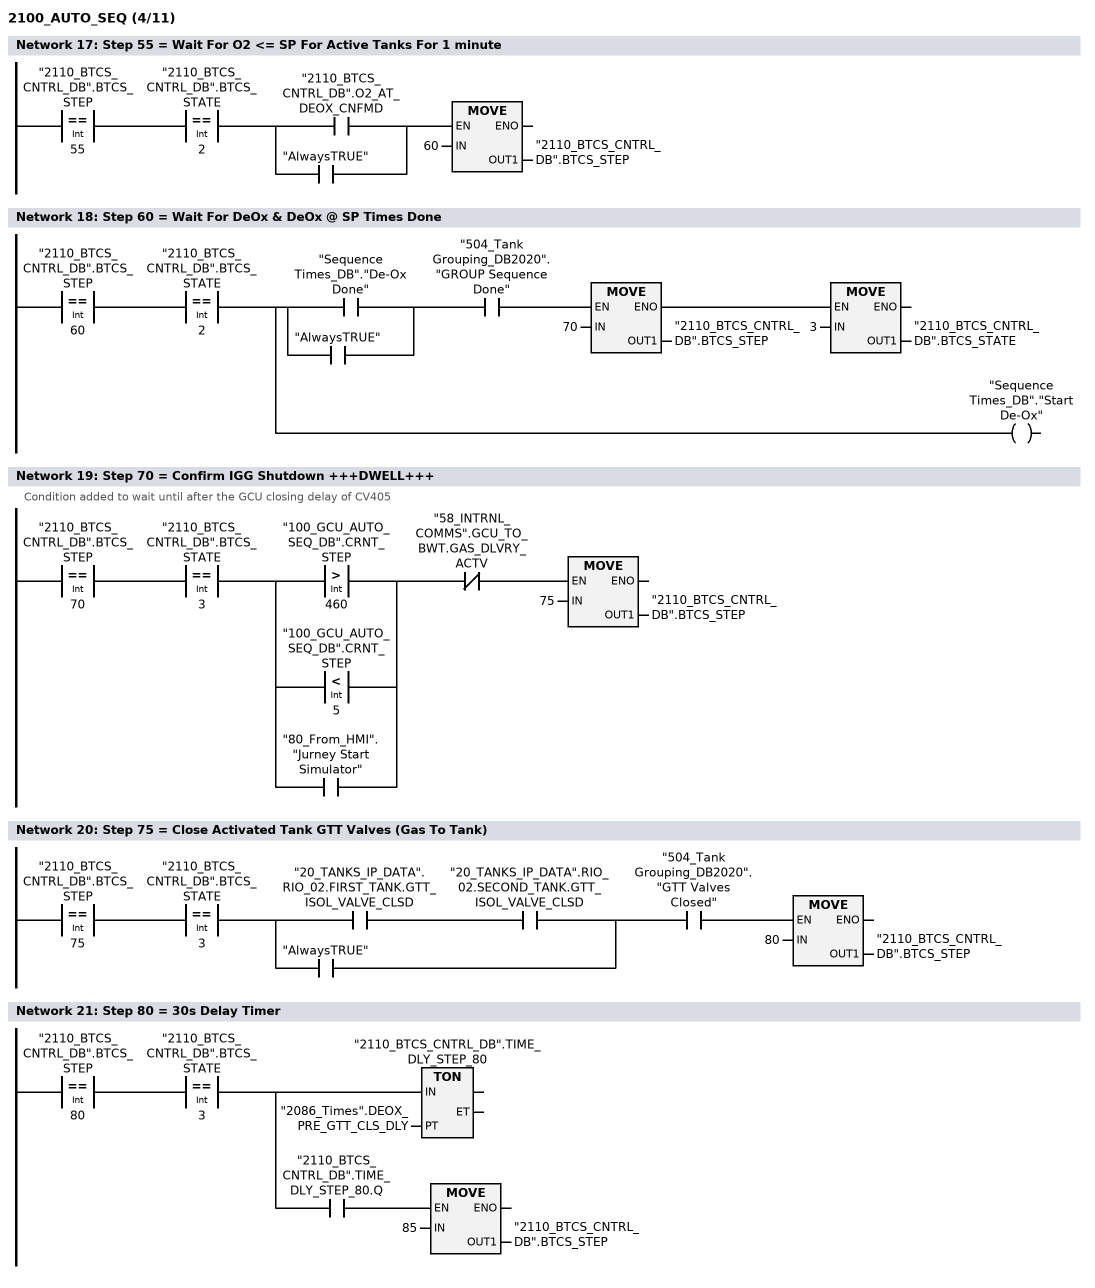
   RUNG wire#powerrail
      { S7_Templates := "SrcType := Int" } EQ_Contact(in1 := "2110_BTCS_CNTRL_DB".BTCS_STEP, in2 := 55)
      { S7_Templates := "SrcType := Int" } EQ_Contact(in1 := "2110_BTCS_CNTRL_DB".BTCS_STATE, in2 := 2)
      wire#w1
      Contact( "2110_BTCS_CNTRL_DB".O2_AT_DEOX_CNFMD )
      wire#w2
      Move(in := 60, out1 => "2110_BTCS_CNTRL_DB".BTCS_STEP)
   END_RUNG
   RUNG wire#w1
      Contact( "AlwaysTRUE" )
   END_RUNG wire#w2
   // the same network as SCL:
   IF ("2110_BTCS_CNTRL_DB".BTCS_STEP = 55) AND ("2110_BTCS_CNTRL_DB".BTCS_STATE = 2) AND ("2110_BTCS_CNTRL_DB".O2_AT_DEOX_CNFMD OR "AlwaysTRUE") THEN
       "2110_BTCS_CNTRL_DB".BTCS_STEP := 60;
   END_IF;
END_REGION

REGION Network 18: Step 60 = Wait For DeOx & DeOx @ SP Times Done
   RUNG wire#powerrail
      { S7_Templates := "SrcType := Int" } EQ_Contact(in1 := "2110_BTCS_CNTRL_DB".BTCS_STEP, in2 := 60)
      { S7_Templates := "SrcType := Int" } EQ_Contact(in1 := "2110_BTCS_CNTRL_DB".BTCS_STATE, in2 := 2)
      wire#w1
      Contact( "Sequence Times_DB"."De-Ox Done" )
      wire#w2
      Contact( "504_Tank Grouping_DB2020"."GROUP Sequence Done" )
      Move(in := 70, out1 => "2110_BTCS_CNTRL_DB".BTCS_STEP)
      Move(in := 3, out1 => "2110_BTCS_CNTRL_DB".BTCS_STATE)
   END_RUNG
   RUNG wire#w1
      Contact( "AlwaysTRUE" )
   END_RUNG wire#w2
   RUNG wire#w1
      Coil( "Sequence Times_DB"."Start De-Ox" )
   END_RUNG
   // the same network as SCL:
   #_w1 := ("2110_BTCS_CNTRL_DB".BTCS_STEP = 60) AND ("2110_BTCS_CNTRL_DB".BTCS_STATE = 2);
   IF #_w1 AND ("Sequence Times_DB"."De-Ox Done" OR "AlwaysTRUE") AND "504_Tank Grouping_DB2020"."GROUP Sequence Done" THEN
       "2110_BTCS_CNTRL_DB".BTCS_STEP := 70;
       "2110_BTCS_CNTRL_DB".BTCS_STATE := 3;
   END_IF;
   "Sequence Times_DB"."Start De-Ox" := #_w1;
END_REGION

REGION Network 19: Step 70 = Confirm IGG Shutdown +++DWELL+++
   // Condition added to wait until after the GCU closing delay of CV405
   RUNG wire#powerrail
      { S7_Templates := "SrcType := Int" } EQ_Contact(in1 := "2110_BTCS_CNTRL_DB".BTCS_STEP, in2 := 70)
      { S7_Templates := "SrcType := Int" } EQ_Contact(in1 := "2110_BTCS_CNTRL_DB".BTCS_STATE, in2 := 3)
      wire#w1
      { S7_Templates := "SrcType := Int" } GT_Contact(in1 := "100_GCU_AUTO_SEQ_DB".CRNT_STEP, in2 := 460)
      wire#w2
      I_Contact( "58_INTRNL_COMMS".GCU_TO_BWT.GAS_DLVRY_ACTV )
      Move(in := 75, out1 => "2110_BTCS_CNTRL_DB".BTCS_STEP)
   END_RUNG
   RUNG wire#w1
      { S7_Templates := "SrcType := Int" } LT_Contact(in1 := "100_GCU_AUTO_SEQ_DB".CRNT_STEP, in2 := 5)
   END_RUNG wire#w2
   RUNG wire#w1
      Contact( "80_From_HMI"."Jurney Start Simulator" )
   END_RUNG wire#w2
   // the same network as SCL:
   IF ("2110_BTCS_CNTRL_DB".BTCS_STEP = 70) AND ("2110_BTCS_CNTRL_DB".BTCS_STATE = 3) AND (("100_GCU_AUTO_SEQ_DB".CRNT_STEP > 460) OR ("100_GCU_AUTO_SEQ_DB".CRNT_STEP < 5) OR "80_From_HMI"."Jurney Start Simulator") AND NOT "58_INTRNL_COMMS".GCU_TO_BWT.GAS_DLVRY_ACTV THEN
       "2110_BTCS_CNTRL_DB".BTCS_STEP := 75;
   END_IF;
END_REGION

REGION Network 20: Step 75 = Close Activated Tank GTT Valves (Gas To Tank)
   RUNG wire#powerrail
      { S7_Templates := "SrcType := Int" } EQ_Contact(in1 := "2110_BTCS_CNTRL_DB".BTCS_STEP, in2 := 75)
      { S7_Templates := "SrcType := Int" } EQ_Contact(in1 := "2110_BTCS_CNTRL_DB".BTCS_STATE, in2 := 3)
      wire#w1
      Contact( "20_TANKS_IP_DATA".RIO_02.FIRST_TANK.GTT_ISOL_VALVE_CLSD )
      Contact( "20_TANKS_IP_DATA".RIO_02.SECOND_TANK.GTT_ISOL_VALVE_CLSD )
      wire#w2
      Contact( "504_Tank Grouping_DB2020"."GTT Valves Closed" )
      Move(in := 80, out1 => "2110_BTCS_CNTRL_DB".BTCS_STEP)
   END_RUNG
   RUNG wire#w1
      Contact( "AlwaysTRUE" )
   END_RUNG wire#w2
   // the same network as SCL:
   IF ("2110_BTCS_CNTRL_DB".BTCS_STEP = 75) AND ("2110_BTCS_CNTRL_DB".BTCS_STATE = 3) AND (("20_TANKS_IP_DATA".RIO_02.FIRST_TANK.GTT_ISOL_VALVE_CLSD AND "20_TANKS_IP_DATA".RIO_02.SECOND_TANK.GTT_ISOL_VALVE_CLSD) OR "AlwaysTRUE") AND "504_Tank Grouping_DB2020"."GTT Valves Closed" THEN
       "2110_BTCS_CNTRL_DB".BTCS_STEP := 80;
   END_IF;
END_REGION

REGION Network 21: Step 80 = 30s Delay Timer
   #_w1 := ("2110_BTCS_CNTRL_DB".BTCS_STEP = 80) AND ("2110_BTCS_CNTRL_DB".BTCS_STATE = 3);
   "2110_BTCS_CNTRL_DB".TIME_DLY_STEP_80.TON(IN := #_w1, PT := "2086_Times".DEOX_PRE_GTT_CLS_DLY);
   IF #_w1 AND "2110_BTCS_CNTRL_DB".TIME_DLY_STEP_80.Q THEN "2110_BTCS_CNTRL_DB".BTCS_STEP := 85; END_IF;
END_REGION

REGION Network 22: Step 85 = Close CV406 Gas to deck valve (Close 406)
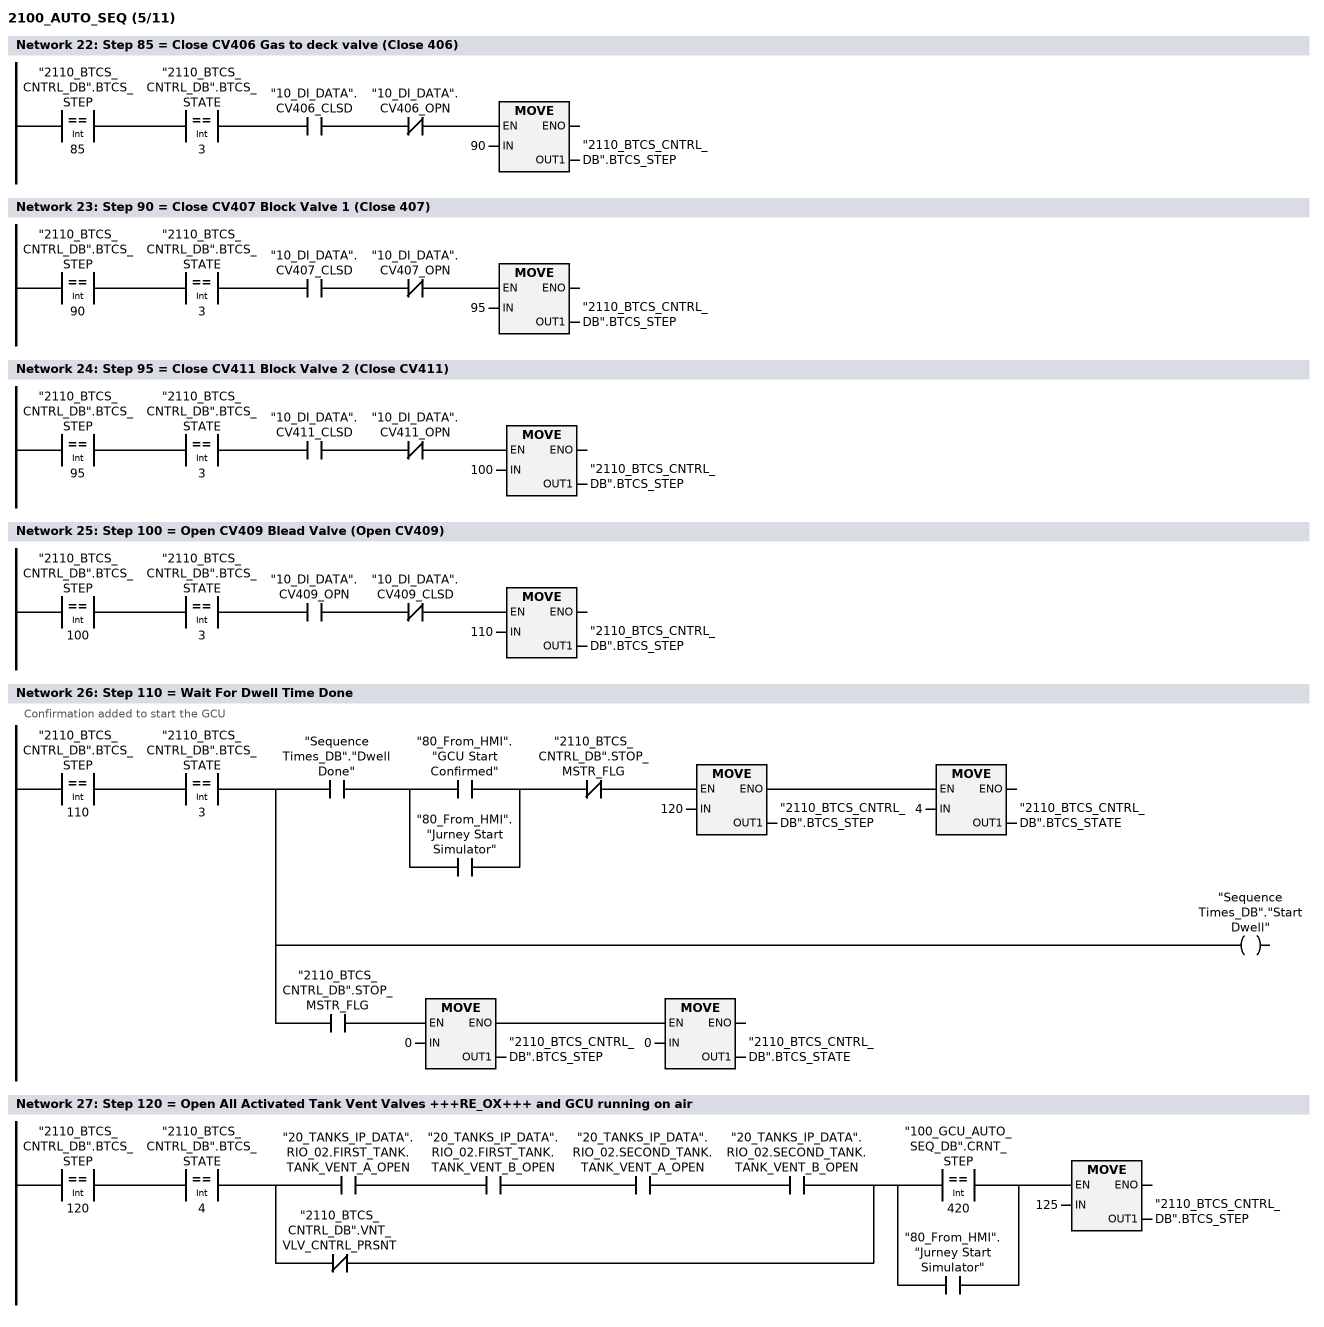
   RUNG wire#powerrail
      { S7_Templates := "SrcType := Int" } EQ_Contact(in1 := "2110_BTCS_CNTRL_DB".BTCS_STEP, in2 := 85)
      { S7_Templates := "SrcType := Int" } EQ_Contact(in1 := "2110_BTCS_CNTRL_DB".BTCS_STATE, in2 := 3)
      Contact( "10_DI_DATA".CV406_CLSD )
      I_Contact( "10_DI_DATA".CV406_OPN )
      Move(in := 90, out1 => "2110_BTCS_CNTRL_DB".BTCS_STEP)
   END_RUNG
   // the same network as SCL:
   IF ("2110_BTCS_CNTRL_DB".BTCS_STEP = 85) AND ("2110_BTCS_CNTRL_DB".BTCS_STATE = 3) AND "10_DI_DATA".CV406_CLSD AND NOT "10_DI_DATA".CV406_OPN THEN
       "2110_BTCS_CNTRL_DB".BTCS_STEP := 90;
   END_IF;
END_REGION

REGION Network 23: Step 90 = Close CV407 Block Valve 1 (Close 407)
   RUNG wire#powerrail
      { S7_Templates := "SrcType := Int" } EQ_Contact(in1 := "2110_BTCS_CNTRL_DB".BTCS_STEP, in2 := 90)
      { S7_Templates := "SrcType := Int" } EQ_Contact(in1 := "2110_BTCS_CNTRL_DB".BTCS_STATE, in2 := 3)
      Contact( "10_DI_DATA".CV407_CLSD )
      I_Contact( "10_DI_DATA".CV407_OPN )
      Move(in := 95, out1 => "2110_BTCS_CNTRL_DB".BTCS_STEP)
   END_RUNG
   // the same network as SCL:
   IF ("2110_BTCS_CNTRL_DB".BTCS_STEP = 90) AND ("2110_BTCS_CNTRL_DB".BTCS_STATE = 3) AND "10_DI_DATA".CV407_CLSD AND NOT "10_DI_DATA".CV407_OPN THEN
       "2110_BTCS_CNTRL_DB".BTCS_STEP := 95;
   END_IF;
END_REGION

REGION Network 24: Step 95 = Close CV411 Block Valve 2 (Close CV411)
   RUNG wire#powerrail
      { S7_Templates := "SrcType := Int" } EQ_Contact(in1 := "2110_BTCS_CNTRL_DB".BTCS_STEP, in2 := 95)
      { S7_Templates := "SrcType := Int" } EQ_Contact(in1 := "2110_BTCS_CNTRL_DB".BTCS_STATE, in2 := 3)
      Contact( "10_DI_DATA".CV411_CLSD )
      I_Contact( "10_DI_DATA".CV411_OPN )
      Move(in := 100, out1 => "2110_BTCS_CNTRL_DB".BTCS_STEP)
   END_RUNG
   // the same network as SCL:
   IF ("2110_BTCS_CNTRL_DB".BTCS_STEP = 95) AND ("2110_BTCS_CNTRL_DB".BTCS_STATE = 3) AND "10_DI_DATA".CV411_CLSD AND NOT "10_DI_DATA".CV411_OPN THEN
       "2110_BTCS_CNTRL_DB".BTCS_STEP := 100;
   END_IF;
END_REGION

REGION Network 25: Step 100 = Open CV409 Blead Valve (Open CV409)
   RUNG wire#powerrail
      { S7_Templates := "SrcType := Int" } EQ_Contact(in1 := "2110_BTCS_CNTRL_DB".BTCS_STEP, in2 := 100)
      { S7_Templates := "SrcType := Int" } EQ_Contact(in1 := "2110_BTCS_CNTRL_DB".BTCS_STATE, in2 := 3)
      Contact( "10_DI_DATA".CV409_OPN )
      I_Contact( "10_DI_DATA".CV409_CLSD )
      Move(in := 110, out1 => "2110_BTCS_CNTRL_DB".BTCS_STEP)
   END_RUNG
   // the same network as SCL:
   IF ("2110_BTCS_CNTRL_DB".BTCS_STEP = 100) AND ("2110_BTCS_CNTRL_DB".BTCS_STATE = 3) AND "10_DI_DATA".CV409_OPN AND NOT "10_DI_DATA".CV409_CLSD THEN
       "2110_BTCS_CNTRL_DB".BTCS_STEP := 110;
   END_IF;
END_REGION

REGION Network 26: Step 110 = Wait For Dwell Time Done
   // Confirmation added to start the GCU
   RUNG wire#powerrail
      { S7_Templates := "SrcType := Int" } EQ_Contact(in1 := "2110_BTCS_CNTRL_DB".BTCS_STEP, in2 := 110)
      { S7_Templates := "SrcType := Int" } EQ_Contact(in1 := "2110_BTCS_CNTRL_DB".BTCS_STATE, in2 := 3)
      wire#w1
      Contact( "Sequence Times_DB"."Dwell Done" )
      wire#w2
      Contact( "80_From_HMI"."GCU Start Confirmed" )
      wire#w3
      I_Contact( "2110_BTCS_CNTRL_DB".STOP_MSTR_FLG )
      Move(in := 120, out1 => "2110_BTCS_CNTRL_DB".BTCS_STEP)
      Move(in := 4, out1 => "2110_BTCS_CNTRL_DB".BTCS_STATE)
   END_RUNG
   RUNG wire#w2
      Contact( "80_From_HMI"."Jurney Start Simulator" )
   END_RUNG wire#w3
   RUNG wire#w1
      Coil( "Sequence Times_DB"."Start Dwell" )
   END_RUNG
   RUNG wire#w1
      Contact( "2110_BTCS_CNTRL_DB".STOP_MSTR_FLG )
      Move(in := 0, out1 => "2110_BTCS_CNTRL_DB".BTCS_STEP)
      Move(in := 0, out1 => "2110_BTCS_CNTRL_DB".BTCS_STATE)
   END_RUNG
   // the same network as SCL:
   #_w1 := ("2110_BTCS_CNTRL_DB".BTCS_STEP = 110) AND ("2110_BTCS_CNTRL_DB".BTCS_STATE = 3);
   IF #_w1 AND "Sequence Times_DB"."Dwell Done" AND ("80_From_HMI"."GCU Start Confirmed" OR "80_From_HMI"."Jurney Start Simulator") AND NOT "2110_BTCS_CNTRL_DB".STOP_MSTR_FLG THEN
       "2110_BTCS_CNTRL_DB".BTCS_STEP := 120;
       "2110_BTCS_CNTRL_DB".BTCS_STATE := 4;
   END_IF;
   "Sequence Times_DB"."Start Dwell" := #_w1;
   IF #_w1 AND "2110_BTCS_CNTRL_DB".STOP_MSTR_FLG THEN
       "2110_BTCS_CNTRL_DB".BTCS_STEP := 0;
       "2110_BTCS_CNTRL_DB".BTCS_STATE := 0;
   END_IF;
END_REGION

REGION Network 27: Step 120 = Open All Activated Tank Vent Valves +++RE_OX+++ and GCU running on air
   RUNG wire#powerrail
      { S7_Templates := "SrcType := Int" } EQ_Contact(in1 := "2110_BTCS_CNTRL_DB".BTCS_STEP, in2 := 120)
      { S7_Templates := "SrcType := Int" } EQ_Contact(in1 := "2110_BTCS_CNTRL_DB".BTCS_STATE, in2 := 4)
      wire#w1
      Contact( "20_TANKS_IP_DATA".RIO_02.FIRST_TANK.TANK_VENT_A_OPEN )
      Contact( "20_TANKS_IP_DATA".RIO_02.FIRST_TANK.TANK_VENT_B_OPEN )
      Contact( "20_TANKS_IP_DATA".RIO_02.SECOND_TANK.TANK_VENT_A_OPEN )
      Contact( "20_TANKS_IP_DATA".RIO_02.SECOND_TANK.TANK_VENT_B_OPEN )
      wire#w2
      { S7_Templates := "SrcType := Int" } EQ_Contact(in1 := "100_GCU_AUTO_SEQ_DB".CRNT_STEP, in2 := 420)
      wire#w3
      Move(in := 125, out1 => "2110_BTCS_CNTRL_DB".BTCS_STEP)
   END_RUNG
   RUNG wire#w1
      I_Contact( "2110_BTCS_CNTRL_DB".VNT_VLV_CNTRL_PRSNT )
   END_RUNG wire#w2
   RUNG wire#w2
      Contact( "80_From_HMI"."Jurney Start Simulator" )
   END_RUNG wire#w3
   // the same network as SCL:
   IF ("2110_BTCS_CNTRL_DB".BTCS_STEP = 120) AND ("2110_BTCS_CNTRL_DB".BTCS_STATE = 4) AND (("20_TANKS_IP_DATA".RIO_02.FIRST_TANK.TANK_VENT_A_OPEN AND "20_TANKS_IP_DATA".RIO_02.FIRST_TANK.TANK_VENT_B_OPEN AND "20_TANKS_IP_DATA".RIO_02.SECOND_TANK.TANK_VENT_A_OPEN AND "20_TANKS_IP_DATA".RIO_02.SECOND_TANK.TANK_VENT_B_OPEN) OR NOT "2110_BTCS_CNTRL_DB".VNT_VLV_CNTRL_PRSNT) AND (("100_GCU_AUTO_SEQ_DB".CRNT_STEP = 420) OR "80_From_HMI"."Jurney Start Simulator") THEN
       "2110_BTCS_CNTRL_DB".BTCS_STEP := 125;
   END_IF;
END_REGION

REGION Network 28: Step 125 = Open CV406 Gas To Deck Valve
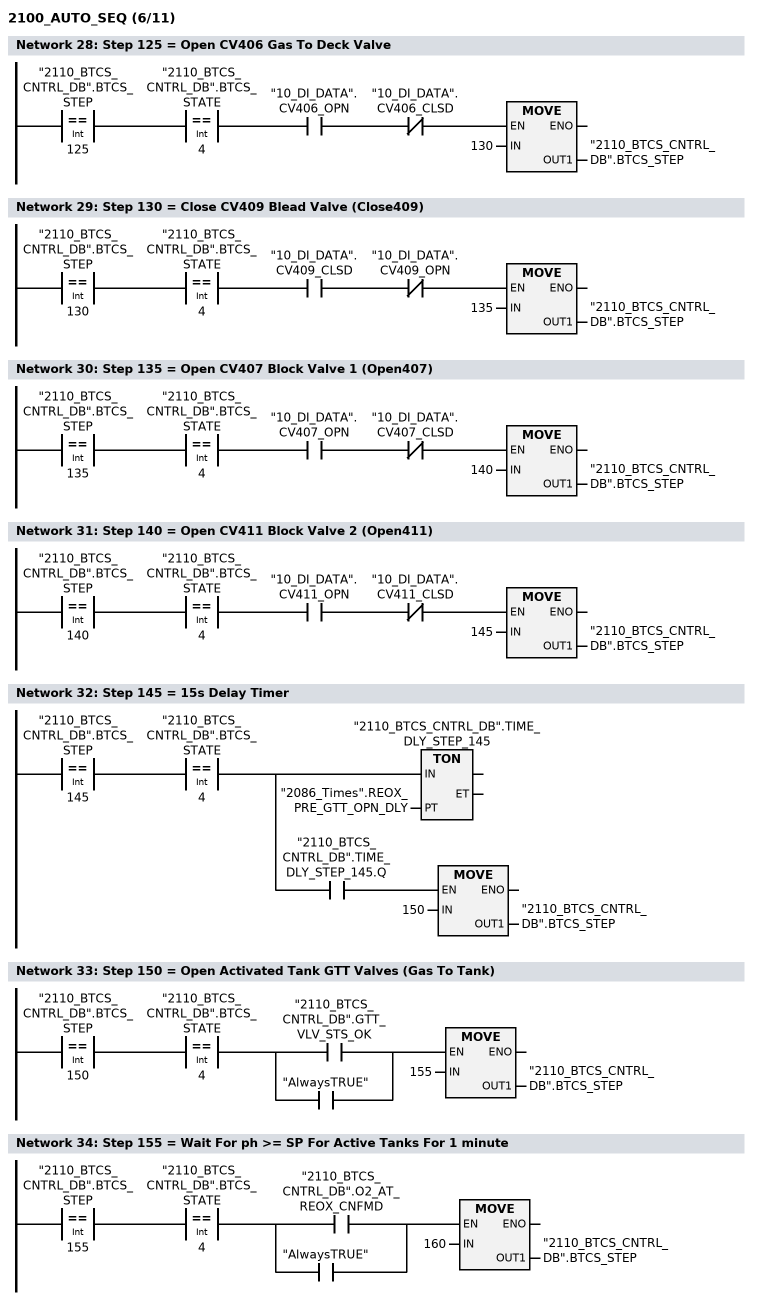
   RUNG wire#powerrail
      { S7_Templates := "SrcType := Int" } EQ_Contact(in1 := "2110_BTCS_CNTRL_DB".BTCS_STEP, in2 := 125)
      { S7_Templates := "SrcType := Int" } EQ_Contact(in1 := "2110_BTCS_CNTRL_DB".BTCS_STATE, in2 := 4)
      Contact( "10_DI_DATA".CV406_OPN )
      I_Contact( "10_DI_DATA".CV406_CLSD )
      Move(in := 130, out1 => "2110_BTCS_CNTRL_DB".BTCS_STEP)
   END_RUNG
   // the same network as SCL:
   IF ("2110_BTCS_CNTRL_DB".BTCS_STEP = 125) AND ("2110_BTCS_CNTRL_DB".BTCS_STATE = 4) AND "10_DI_DATA".CV406_OPN AND NOT "10_DI_DATA".CV406_CLSD THEN
       "2110_BTCS_CNTRL_DB".BTCS_STEP := 130;
   END_IF;
END_REGION

REGION Network 29: Step 130 = Close CV409 Blead Valve (Close409)
   RUNG wire#powerrail
      { S7_Templates := "SrcType := Int" } EQ_Contact(in1 := "2110_BTCS_CNTRL_DB".BTCS_STEP, in2 := 130)
      { S7_Templates := "SrcType := Int" } EQ_Contact(in1 := "2110_BTCS_CNTRL_DB".BTCS_STATE, in2 := 4)
      Contact( "10_DI_DATA".CV409_CLSD )
      I_Contact( "10_DI_DATA".CV409_OPN )
      Move(in := 135, out1 => "2110_BTCS_CNTRL_DB".BTCS_STEP)
   END_RUNG
   // the same network as SCL:
   IF ("2110_BTCS_CNTRL_DB".BTCS_STEP = 130) AND ("2110_BTCS_CNTRL_DB".BTCS_STATE = 4) AND "10_DI_DATA".CV409_CLSD AND NOT "10_DI_DATA".CV409_OPN THEN
       "2110_BTCS_CNTRL_DB".BTCS_STEP := 135;
   END_IF;
END_REGION

REGION Network 30: Step 135 = Open CV407 Block Valve 1 (Open407)
   RUNG wire#powerrail
      { S7_Templates := "SrcType := Int" } EQ_Contact(in1 := "2110_BTCS_CNTRL_DB".BTCS_STEP, in2 := 135)
      { S7_Templates := "SrcType := Int" } EQ_Contact(in1 := "2110_BTCS_CNTRL_DB".BTCS_STATE, in2 := 4)
      Contact( "10_DI_DATA".CV407_OPN )
      I_Contact( "10_DI_DATA".CV407_CLSD )
      Move(in := 140, out1 => "2110_BTCS_CNTRL_DB".BTCS_STEP)
   END_RUNG
   // the same network as SCL:
   IF ("2110_BTCS_CNTRL_DB".BTCS_STEP = 135) AND ("2110_BTCS_CNTRL_DB".BTCS_STATE = 4) AND "10_DI_DATA".CV407_OPN AND NOT "10_DI_DATA".CV407_CLSD THEN
       "2110_BTCS_CNTRL_DB".BTCS_STEP := 140;
   END_IF;
END_REGION

REGION Network 31: Step 140 = Open CV411 Block Valve 2 (Open411)
   RUNG wire#powerrail
      { S7_Templates := "SrcType := Int" } EQ_Contact(in1 := "2110_BTCS_CNTRL_DB".BTCS_STEP, in2 := 140)
      { S7_Templates := "SrcType := Int" } EQ_Contact(in1 := "2110_BTCS_CNTRL_DB".BTCS_STATE, in2 := 4)
      Contact( "10_DI_DATA".CV411_OPN )
      I_Contact( "10_DI_DATA".CV411_CLSD )
      Move(in := 145, out1 => "2110_BTCS_CNTRL_DB".BTCS_STEP)
   END_RUNG
   // the same network as SCL:
   IF ("2110_BTCS_CNTRL_DB".BTCS_STEP = 140) AND ("2110_BTCS_CNTRL_DB".BTCS_STATE = 4) AND "10_DI_DATA".CV411_OPN AND NOT "10_DI_DATA".CV411_CLSD THEN
       "2110_BTCS_CNTRL_DB".BTCS_STEP := 145;
   END_IF;
END_REGION

REGION Network 32: Step 145 = 15s Delay Timer
   #_w1 := ("2110_BTCS_CNTRL_DB".BTCS_STEP = 145) AND ("2110_BTCS_CNTRL_DB".BTCS_STATE = 4);
   "2110_BTCS_CNTRL_DB".TIME_DLY_STEP_145.TON(IN := #_w1, PT := "2086_Times".REOX_PRE_GTT_OPN_DLY);
   IF #_w1 AND "2110_BTCS_CNTRL_DB".TIME_DLY_STEP_145.Q THEN "2110_BTCS_CNTRL_DB".BTCS_STEP := 150; END_IF;
END_REGION

REGION Network 33: Step 150 = Open Activated Tank GTT Valves (Gas To Tank)
   RUNG wire#powerrail
      { S7_Templates := "SrcType := Int" } EQ_Contact(in1 := "2110_BTCS_CNTRL_DB".BTCS_STEP, in2 := 150)
      { S7_Templates := "SrcType := Int" } EQ_Contact(in1 := "2110_BTCS_CNTRL_DB".BTCS_STATE, in2 := 4)
      wire#w1
      Contact( "2110_BTCS_CNTRL_DB".GTT_VLV_STS_OK )
      wire#w2
      Move(in := 155, out1 => "2110_BTCS_CNTRL_DB".BTCS_STEP)
   END_RUNG
   RUNG wire#w1
      Contact( "AlwaysTRUE" )
   END_RUNG wire#w2
   // the same network as SCL:
   IF ("2110_BTCS_CNTRL_DB".BTCS_STEP = 150) AND ("2110_BTCS_CNTRL_DB".BTCS_STATE = 4) AND ("2110_BTCS_CNTRL_DB".GTT_VLV_STS_OK OR "AlwaysTRUE") THEN
       "2110_BTCS_CNTRL_DB".BTCS_STEP := 155;
   END_IF;
END_REGION

REGION Network 34: Step 155 = Wait For ph >= SP For Active Tanks For 1 minute
   RUNG wire#powerrail
      { S7_Templates := "SrcType := Int" } EQ_Contact(in1 := "2110_BTCS_CNTRL_DB".BTCS_STEP, in2 := 155)
      { S7_Templates := "SrcType := Int" } EQ_Contact(in1 := "2110_BTCS_CNTRL_DB".BTCS_STATE, in2 := 4)
      wire#w1
      Contact( "2110_BTCS_CNTRL_DB".O2_AT_REOX_CNFMD )
      wire#w2
      Move(in := 160, out1 => "2110_BTCS_CNTRL_DB".BTCS_STEP)
   END_RUNG
   RUNG wire#w1
      Contact( "AlwaysTRUE" )
   END_RUNG wire#w2
   // the same network as SCL:
   IF ("2110_BTCS_CNTRL_DB".BTCS_STEP = 155) AND ("2110_BTCS_CNTRL_DB".BTCS_STATE = 4) AND ("2110_BTCS_CNTRL_DB".O2_AT_REOX_CNFMD OR "AlwaysTRUE") THEN
       "2110_BTCS_CNTRL_DB".BTCS_STEP := 160;
   END_IF;
END_REGION

REGION Network 35: Step 160 = Wait For ReOx & ReOx @ SP Times Done
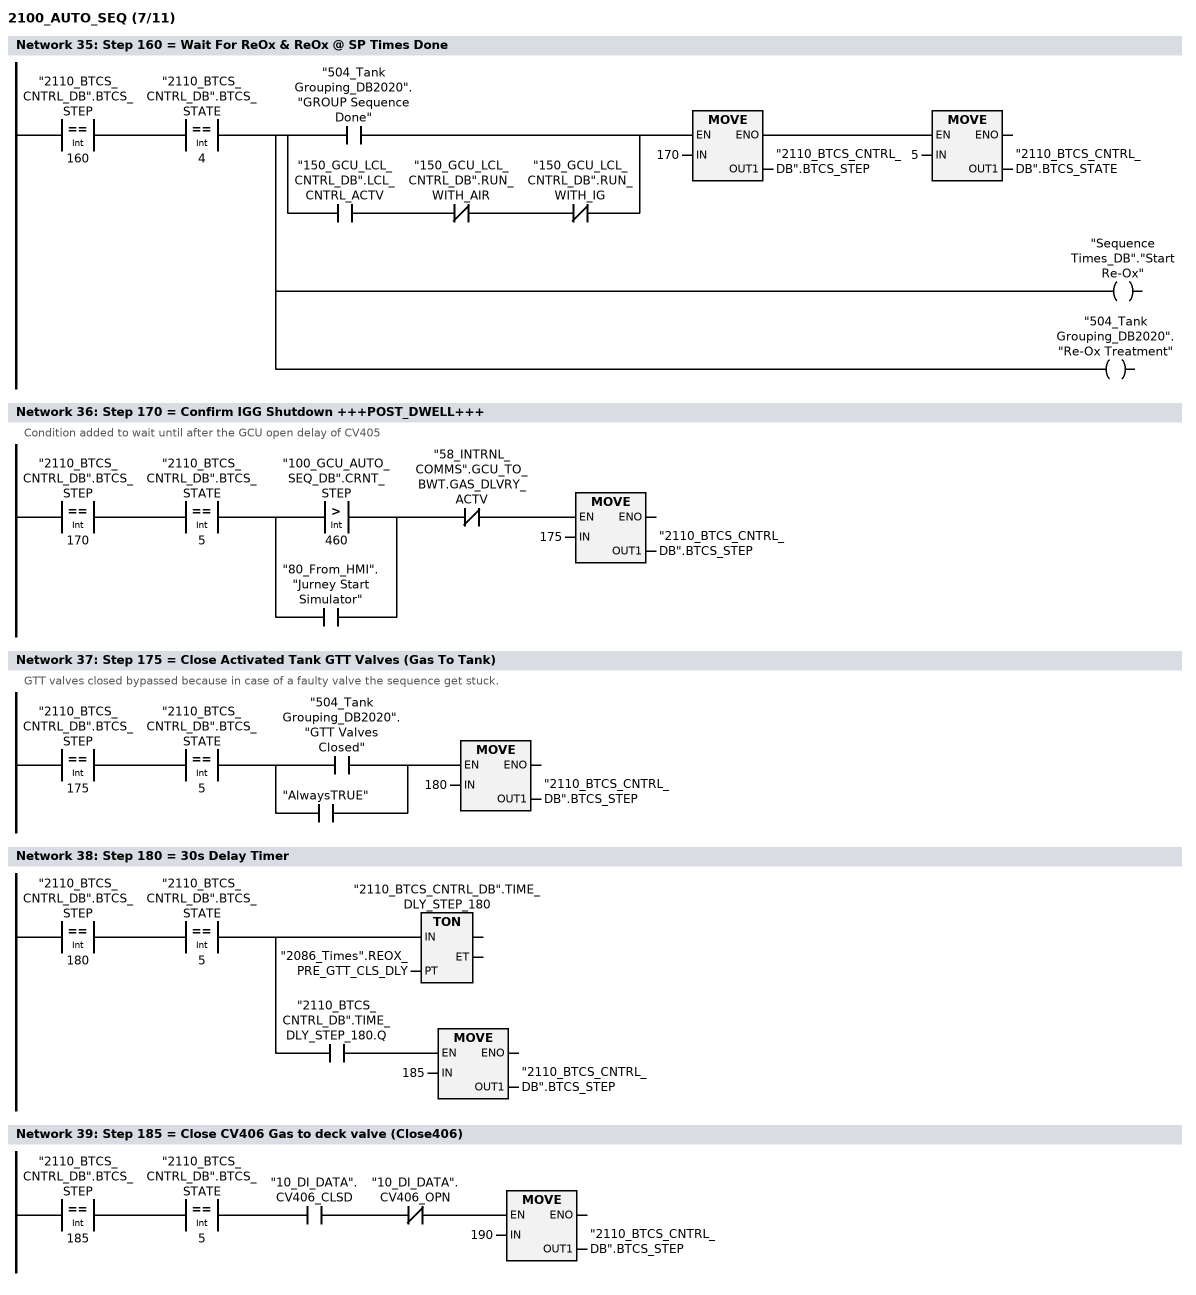
   RUNG wire#powerrail
      { S7_Templates := "SrcType := Int" } EQ_Contact(in1 := "2110_BTCS_CNTRL_DB".BTCS_STEP, in2 := 160)
      { S7_Templates := "SrcType := Int" } EQ_Contact(in1 := "2110_BTCS_CNTRL_DB".BTCS_STATE, in2 := 4)
      wire#w1
      Contact( "504_Tank Grouping_DB2020"."GROUP Sequence Done" )
      wire#w2
      Move(in := 170, out1 => "2110_BTCS_CNTRL_DB".BTCS_STEP)
      Move(in := 5, out1 => "2110_BTCS_CNTRL_DB".BTCS_STATE)
   END_RUNG
   RUNG wire#w1
      Contact( "150_GCU_LCL_CNTRL_DB".LCL_CNTRL_ACTV )
      I_Contact( "150_GCU_LCL_CNTRL_DB".RUN_WITH_AIR )
      I_Contact( "150_GCU_LCL_CNTRL_DB".RUN_WITH_IG )
   END_RUNG wire#w2
   RUNG wire#w1
      Coil( "Sequence Times_DB"."Start Re-Ox" )
   END_RUNG
   RUNG wire#w1
      Coil( "504_Tank Grouping_DB2020"."Re-Ox Treatment" )
   END_RUNG
   // the same network as SCL:
   #_w1 := ("2110_BTCS_CNTRL_DB".BTCS_STEP = 160) AND ("2110_BTCS_CNTRL_DB".BTCS_STATE = 4);
   IF #_w1 AND ("504_Tank Grouping_DB2020"."GROUP Sequence Done" OR ("150_GCU_LCL_CNTRL_DB".LCL_CNTRL_ACTV AND NOT "150_GCU_LCL_CNTRL_DB".RUN_WITH_AIR AND NOT "150_GCU_LCL_CNTRL_DB".RUN_WITH_IG)) THEN
       "2110_BTCS_CNTRL_DB".BTCS_STEP := 170;
       "2110_BTCS_CNTRL_DB".BTCS_STATE := 5;
   END_IF;
   "Sequence Times_DB"."Start Re-Ox" := #_w1;
   "504_Tank Grouping_DB2020"."Re-Ox Treatment" := #_w1;
END_REGION

REGION Network 36: Step 170 = Confirm IGG Shutdown +++POST_DWELL+++
   // Condition added to wait until after the GCU open delay of CV405
   RUNG wire#powerrail
      { S7_Templates := "SrcType := Int" } EQ_Contact(in1 := "2110_BTCS_CNTRL_DB".BTCS_STEP, in2 := 170)
      { S7_Templates := "SrcType := Int" } EQ_Contact(in1 := "2110_BTCS_CNTRL_DB".BTCS_STATE, in2 := 5)
      wire#w1
      { S7_Templates := "SrcType := Int" } GT_Contact(in1 := "100_GCU_AUTO_SEQ_DB".CRNT_STEP, in2 := 460)
      wire#w2
      I_Contact( "58_INTRNL_COMMS".GCU_TO_BWT.GAS_DLVRY_ACTV )
      Move(in := 175, out1 => "2110_BTCS_CNTRL_DB".BTCS_STEP)
   END_RUNG
   RUNG wire#w1
      Contact( "80_From_HMI"."Jurney Start Simulator" )
   END_RUNG wire#w2
   // the same network as SCL:
   IF ("2110_BTCS_CNTRL_DB".BTCS_STEP = 170) AND ("2110_BTCS_CNTRL_DB".BTCS_STATE = 5) AND (("100_GCU_AUTO_SEQ_DB".CRNT_STEP > 460) OR "80_From_HMI"."Jurney Start Simulator") AND NOT "58_INTRNL_COMMS".GCU_TO_BWT.GAS_DLVRY_ACTV THEN
       "2110_BTCS_CNTRL_DB".BTCS_STEP := 175;
   END_IF;
END_REGION

REGION Network 37: Step 175 = Close Activated Tank GTT Valves (Gas To Tank)
   // GTT valves closed bypassed because in case of a faulty valve the sequence get stuck.
   RUNG wire#powerrail
      { S7_Templates := "SrcType := Int" } EQ_Contact(in1 := "2110_BTCS_CNTRL_DB".BTCS_STEP, in2 := 175)
      { S7_Templates := "SrcType := Int" } EQ_Contact(in1 := "2110_BTCS_CNTRL_DB".BTCS_STATE, in2 := 5)
      wire#w1
      Contact( "504_Tank Grouping_DB2020"."GTT Valves Closed" )
      wire#w2
      Move(in := 180, out1 => "2110_BTCS_CNTRL_DB".BTCS_STEP)
   END_RUNG
   RUNG wire#w1
      Contact( "AlwaysTRUE" )
   END_RUNG wire#w2
   // the same network as SCL:
   IF ("2110_BTCS_CNTRL_DB".BTCS_STEP = 175) AND ("2110_BTCS_CNTRL_DB".BTCS_STATE = 5) AND ("504_Tank Grouping_DB2020"."GTT Valves Closed" OR "AlwaysTRUE") THEN
       "2110_BTCS_CNTRL_DB".BTCS_STEP := 180;
   END_IF;
END_REGION

REGION Network 38: Step 180 = 30s Delay Timer
   #_w1 := ("2110_BTCS_CNTRL_DB".BTCS_STEP = 180) AND ("2110_BTCS_CNTRL_DB".BTCS_STATE = 5);
   "2110_BTCS_CNTRL_DB".TIME_DLY_STEP_180.TON(IN := #_w1, PT := "2086_Times".REOX_PRE_GTT_CLS_DLY);
   IF #_w1 AND "2110_BTCS_CNTRL_DB".TIME_DLY_STEP_180.Q THEN "2110_BTCS_CNTRL_DB".BTCS_STEP := 185; END_IF;
END_REGION

REGION Network 39: Step 185 = Close CV406 Gas to deck valve (Close406)
   RUNG wire#powerrail
      { S7_Templates := "SrcType := Int" } EQ_Contact(in1 := "2110_BTCS_CNTRL_DB".BTCS_STEP, in2 := 185)
      { S7_Templates := "SrcType := Int" } EQ_Contact(in1 := "2110_BTCS_CNTRL_DB".BTCS_STATE, in2 := 5)
      Contact( "10_DI_DATA".CV406_CLSD )
      I_Contact( "10_DI_DATA".CV406_OPN )
      Move(in := 190, out1 => "2110_BTCS_CNTRL_DB".BTCS_STEP)
   END_RUNG
   // the same network as SCL:
   IF ("2110_BTCS_CNTRL_DB".BTCS_STEP = 185) AND ("2110_BTCS_CNTRL_DB".BTCS_STATE = 5) AND "10_DI_DATA".CV406_CLSD AND NOT "10_DI_DATA".CV406_OPN THEN
       "2110_BTCS_CNTRL_DB".BTCS_STEP := 190;
   END_IF;
END_REGION

REGION Network 40: Step 190 = Close CV407 Block Valve 1 (Close CV407)
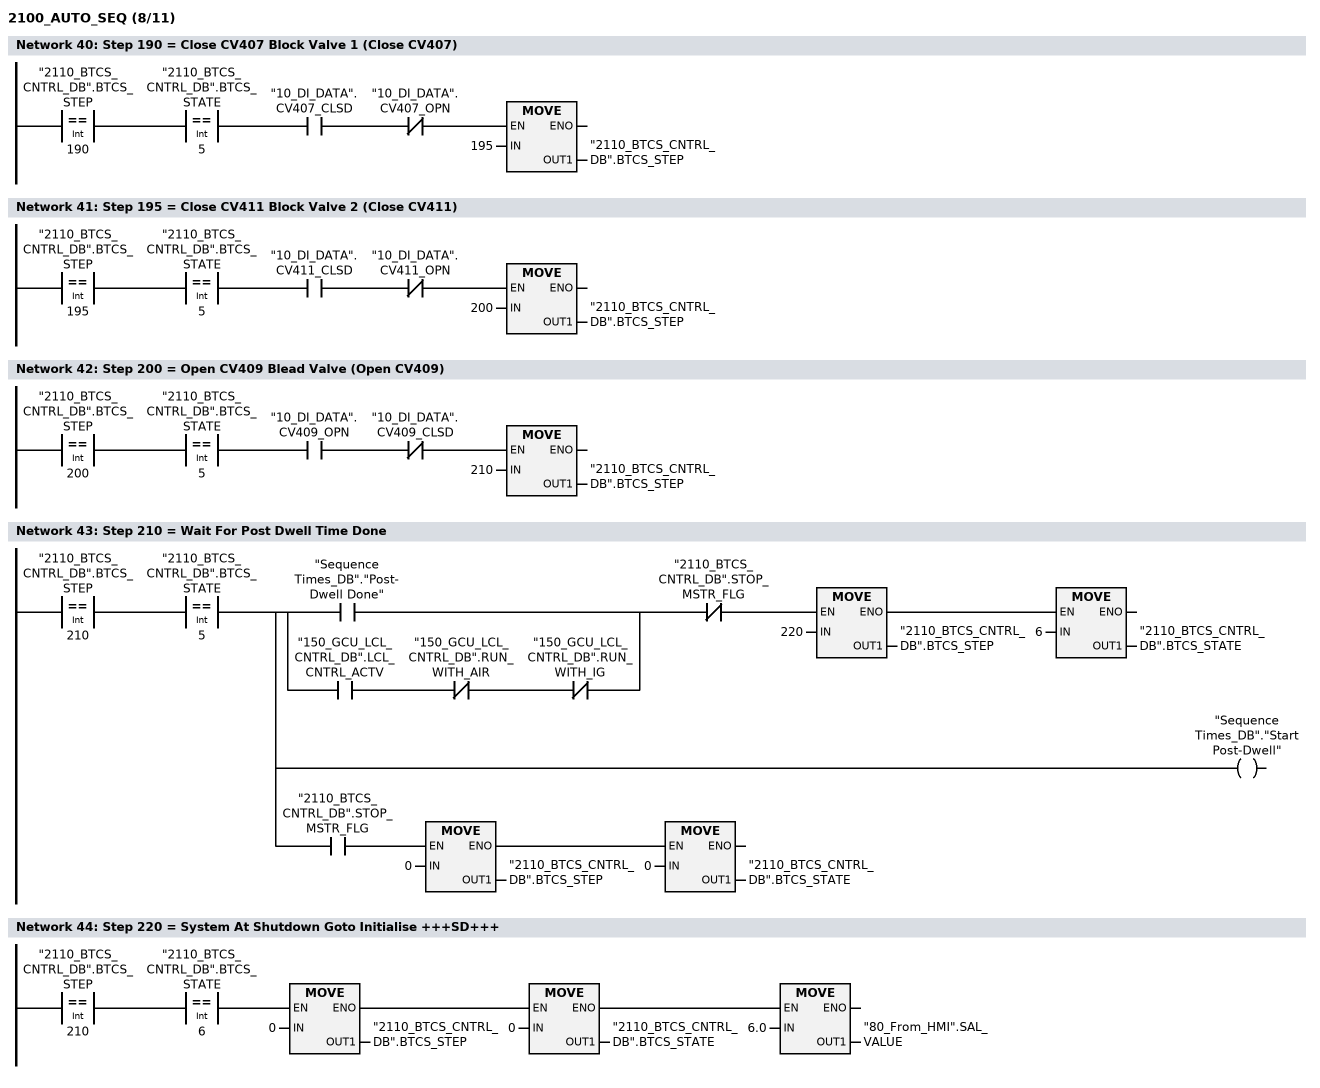
   RUNG wire#powerrail
      { S7_Templates := "SrcType := Int" } EQ_Contact(in1 := "2110_BTCS_CNTRL_DB".BTCS_STEP, in2 := 190)
      { S7_Templates := "SrcType := Int" } EQ_Contact(in1 := "2110_BTCS_CNTRL_DB".BTCS_STATE, in2 := 5)
      Contact( "10_DI_DATA".CV407_CLSD )
      I_Contact( "10_DI_DATA".CV407_OPN )
      Move(in := 195, out1 => "2110_BTCS_CNTRL_DB".BTCS_STEP)
   END_RUNG
   // the same network as SCL:
   IF ("2110_BTCS_CNTRL_DB".BTCS_STEP = 190) AND ("2110_BTCS_CNTRL_DB".BTCS_STATE = 5) AND "10_DI_DATA".CV407_CLSD AND NOT "10_DI_DATA".CV407_OPN THEN
       "2110_BTCS_CNTRL_DB".BTCS_STEP := 195;
   END_IF;
END_REGION

REGION Network 41: Step 195 = Close CV411 Block Valve 2 (Close CV411)
   RUNG wire#powerrail
      { S7_Templates := "SrcType := Int" } EQ_Contact(in1 := "2110_BTCS_CNTRL_DB".BTCS_STEP, in2 := 195)
      { S7_Templates := "SrcType := Int" } EQ_Contact(in1 := "2110_BTCS_CNTRL_DB".BTCS_STATE, in2 := 5)
      Contact( "10_DI_DATA".CV411_CLSD )
      I_Contact( "10_DI_DATA".CV411_OPN )
      Move(in := 200, out1 => "2110_BTCS_CNTRL_DB".BTCS_STEP)
   END_RUNG
   // the same network as SCL:
   IF ("2110_BTCS_CNTRL_DB".BTCS_STEP = 195) AND ("2110_BTCS_CNTRL_DB".BTCS_STATE = 5) AND "10_DI_DATA".CV411_CLSD AND NOT "10_DI_DATA".CV411_OPN THEN
       "2110_BTCS_CNTRL_DB".BTCS_STEP := 200;
   END_IF;
END_REGION

REGION Network 42: Step 200 = Open CV409 Blead Valve (Open CV409)
   RUNG wire#powerrail
      { S7_Templates := "SrcType := Int" } EQ_Contact(in1 := "2110_BTCS_CNTRL_DB".BTCS_STEP, in2 := 200)
      { S7_Templates := "SrcType := Int" } EQ_Contact(in1 := "2110_BTCS_CNTRL_DB".BTCS_STATE, in2 := 5)
      Contact( "10_DI_DATA".CV409_OPN )
      I_Contact( "10_DI_DATA".CV409_CLSD )
      Move(in := 210, out1 => "2110_BTCS_CNTRL_DB".BTCS_STEP)
   END_RUNG
   // the same network as SCL:
   IF ("2110_BTCS_CNTRL_DB".BTCS_STEP = 200) AND ("2110_BTCS_CNTRL_DB".BTCS_STATE = 5) AND "10_DI_DATA".CV409_OPN AND NOT "10_DI_DATA".CV409_CLSD THEN
       "2110_BTCS_CNTRL_DB".BTCS_STEP := 210;
   END_IF;
END_REGION

REGION Network 43: Step 210 = Wait For Post Dwell Time Done
   RUNG wire#powerrail
      { S7_Templates := "SrcType := Int" } EQ_Contact(in1 := "2110_BTCS_CNTRL_DB".BTCS_STEP, in2 := 210)
      { S7_Templates := "SrcType := Int" } EQ_Contact(in1 := "2110_BTCS_CNTRL_DB".BTCS_STATE, in2 := 5)
      wire#w1
      Contact( "Sequence Times_DB"."Post-Dwell Done" )
      wire#w2
      I_Contact( "2110_BTCS_CNTRL_DB".STOP_MSTR_FLG )
      Move(in := 220, out1 => "2110_BTCS_CNTRL_DB".BTCS_STEP)
      Move(in := 6, out1 => "2110_BTCS_CNTRL_DB".BTCS_STATE)
   END_RUNG
   RUNG wire#w1
      Contact( "150_GCU_LCL_CNTRL_DB".LCL_CNTRL_ACTV )
      I_Contact( "150_GCU_LCL_CNTRL_DB".RUN_WITH_AIR )
      I_Contact( "150_GCU_LCL_CNTRL_DB".RUN_WITH_IG )
   END_RUNG wire#w2
   RUNG wire#w1
      Coil( "Sequence Times_DB"."Start Post-Dwell" )
   END_RUNG
   RUNG wire#w1
      Contact( "2110_BTCS_CNTRL_DB".STOP_MSTR_FLG )
      Move(in := 0, out1 => "2110_BTCS_CNTRL_DB".BTCS_STEP)
      Move(in := 0, out1 => "2110_BTCS_CNTRL_DB".BTCS_STATE)
   END_RUNG
   // the same network as SCL:
   #_w1 := ("2110_BTCS_CNTRL_DB".BTCS_STEP = 210) AND ("2110_BTCS_CNTRL_DB".BTCS_STATE = 5);
   IF #_w1 AND ("Sequence Times_DB"."Post-Dwell Done" OR ("150_GCU_LCL_CNTRL_DB".LCL_CNTRL_ACTV AND NOT "150_GCU_LCL_CNTRL_DB".RUN_WITH_AIR AND NOT "150_GCU_LCL_CNTRL_DB".RUN_WITH_IG)) AND NOT "2110_BTCS_CNTRL_DB".STOP_MSTR_FLG THEN
       "2110_BTCS_CNTRL_DB".BTCS_STEP := 220;
       "2110_BTCS_CNTRL_DB".BTCS_STATE := 6;
   END_IF;
   "Sequence Times_DB"."Start Post-Dwell" := #_w1;
   IF #_w1 AND "2110_BTCS_CNTRL_DB".STOP_MSTR_FLG THEN
       "2110_BTCS_CNTRL_DB".BTCS_STEP := 0;
       "2110_BTCS_CNTRL_DB".BTCS_STATE := 0;
   END_IF;
END_REGION

REGION Network 44: Step 220 = System At Shutdown Goto Initialise +++SD+++
   RUNG wire#powerrail
      { S7_Templates := "SrcType := Int" } EQ_Contact(in1 := "2110_BTCS_CNTRL_DB".BTCS_STEP, in2 := 210)
      { S7_Templates := "SrcType := Int" } EQ_Contact(in1 := "2110_BTCS_CNTRL_DB".BTCS_STATE, in2 := 6)
      Move(in := 0, out1 => "2110_BTCS_CNTRL_DB".BTCS_STEP)
      Move(in := 0, out1 => "2110_BTCS_CNTRL_DB".BTCS_STATE)
      Move(in := 6.0, out1 => "80_From_HMI".SAL_VALUE)
   END_RUNG
   // the same network as SCL:
   #_w1 := ("2110_BTCS_CNTRL_DB".BTCS_STEP = 210) AND ("2110_BTCS_CNTRL_DB".BTCS_STATE = 6);
   IF #_w1 THEN
       "2110_BTCS_CNTRL_DB".BTCS_STEP := 0;
       "2110_BTCS_CNTRL_DB".BTCS_STATE := 0;
       "80_From_HMI".SAL_VALUE := 6.0;
   END_IF;
END_REGION

REGION Network 46: Sequence Times